(* Logix 5000 project; controller FV vendor 1 type 14 code 217 rev 31.11; software revision 31.00; part 33 of 63 *)
(* tags used below, declared in another part *)
   Alarm_Reset : BOOL;
   CheckTimeMask : INT;
   CLOCK_system_set : BOOL;
   CLOCKsetvalues : DINT[7];
   CurrentTime : DateTime;
   CWD : CHECKWORD_FLAGS;
   FR_data_file_value_to_move : DINT;
   FR_dow_addon_tag : DayOfWeek;
   FR_dow_timer : TIMER;
   FR_N120 : INT[265];   // YEAST CROP Yeast Cropping Main
   FR_N160 : INT[265];   // VESSEL Vessel Working Direc tory
   FR_N255 : INT[265];   // CHECKWORDS
   FR_N99 : INT[265];   // COMMENT Comment Lines
   FR_PANELESTOP : PlantItem;   // PANELESTOP
   FR_PILZ : PlantItem;   // PILZ
   FR_SFile : INT[255];   // SLC Equivalent System File, So Original Code Can Remain
   FR_T121 : TIMER[255];   // YEAST CROP
   FtoF_raw_input : REAL;
   FV_SFile : INT[255];   // SLC Equivalent System File, So Original Code Can Remain
   ItoF_raw_input : INT;
   One_Second_One_Scan : ALIAS FOR One_Second_1_scan;
   scale_analog_int : DINT;
   scale_analog_result : REAL;
   scale_eu_max : REAL;
   scale_eu_min : REAL;
   scale_raw_input : REAL;
   scale_raw_max : REAL;
   scale_raw_min : REAL;
   scale_routine_active : BOOL;
   scale_temp : REAL;
(* FR_Common, continued *)

ROUTINE FR_YEAST_ST_120   (* ladder *)
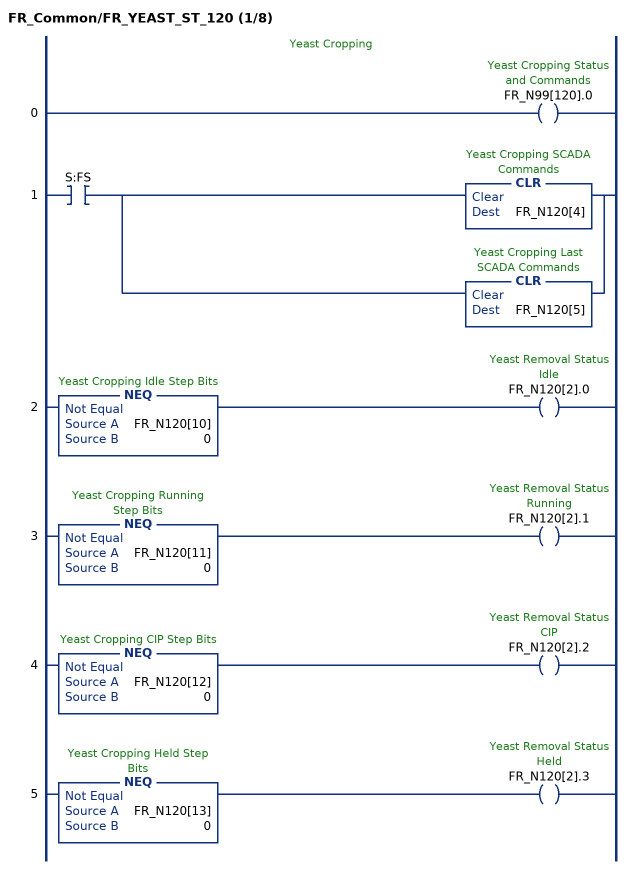
   // Yeast Cropping
   0: OTE(FR_N99[120].0);
   1: XIC(S:FS)[CLR(FR_N120[4]) ,CLR(FR_N120[5]) ];
   2: NEQ(FR_N120[10],0)OTE(FR_N120[2].0);
   3: NEQ(FR_N120[11],0)OTE(FR_N120[2].1);
   4: NEQ(FR_N120[12],0)OTE(FR_N120[2].2);
   5: NEQ(FR_N120[13],0)OTE(FR_N120[2].3);
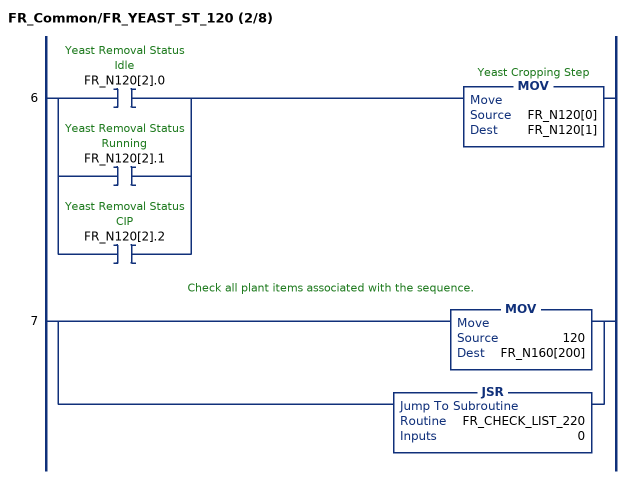
   6: [XIC(FR_N120[2].0) ,XIC(FR_N120[2].1) ,XIC(FR_N120[2].2) ]MOV(FR_N120[0],FR_N120[1]);
   // Check all plant items associated with the sequence.
   7: [MOV(120,FR_N160[200]) ,JSR(FR_CHECK_LIST_220,0) ];
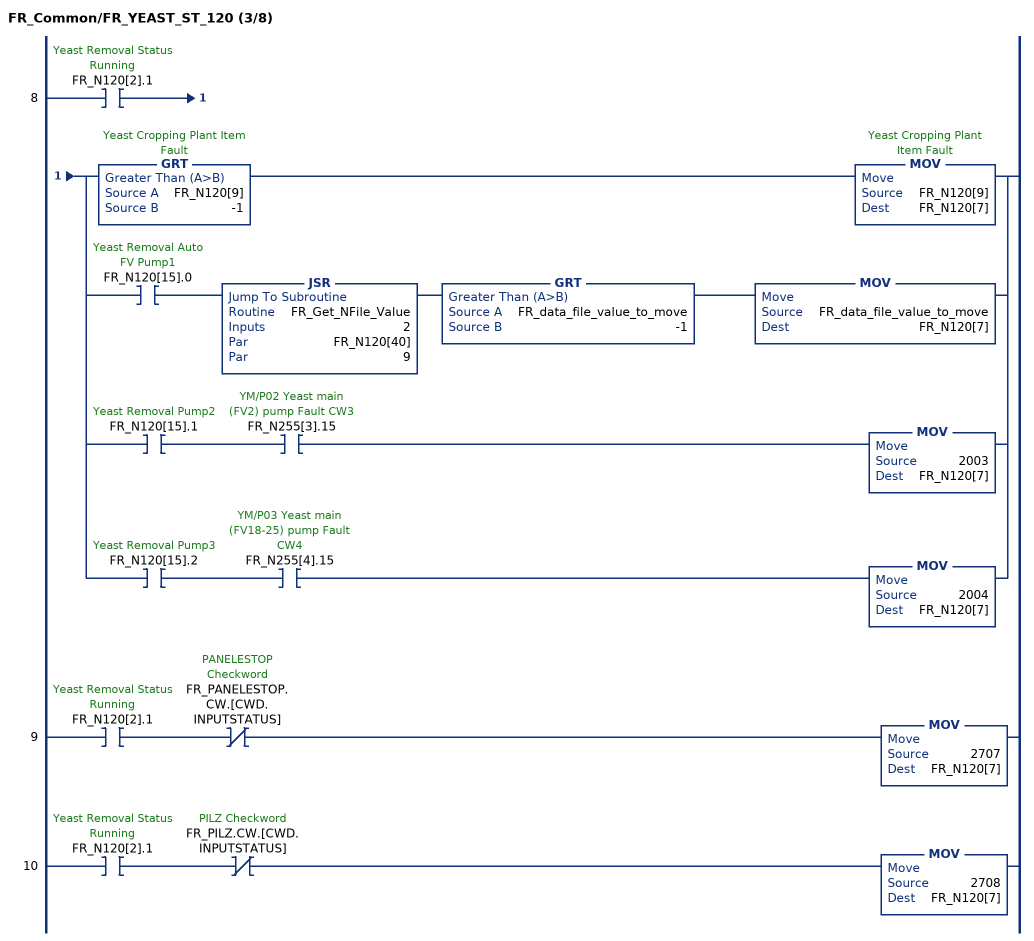
   8: XIC(FR_N120[2].1)[GRT(FR_N120[9],-1) MOV(FR_N120[9],FR_N120[7]) ,XIC(FR_N120[15].0) JSR(FR_Get_NFile_Value,2,FR_N120[40],9) GRT(FR_data_file_value_to_move,-1) MOV(FR_data_file_value_to_move,FR_N120[7]) ,XIC(FR_N120[15].1) XIC(FR_N255[3].15) MOV(2003,FR_N120[7]) ,XIC(FR_N120[15].2) XIC(FR_N255[4].15) MOV(2004,FR_N120[7]) ];
   9: XIC(FR_N120[2].1)XIO(FR_PANELESTOP.CW.[CWD.INPUTSTATUS])MOV(2707,FR_N120[7]);
   10: XIC(FR_N120[2].1)XIO(FR_PILZ.CW.[CWD.INPUTSTATUS])MOV(2708,FR_N120[7]);
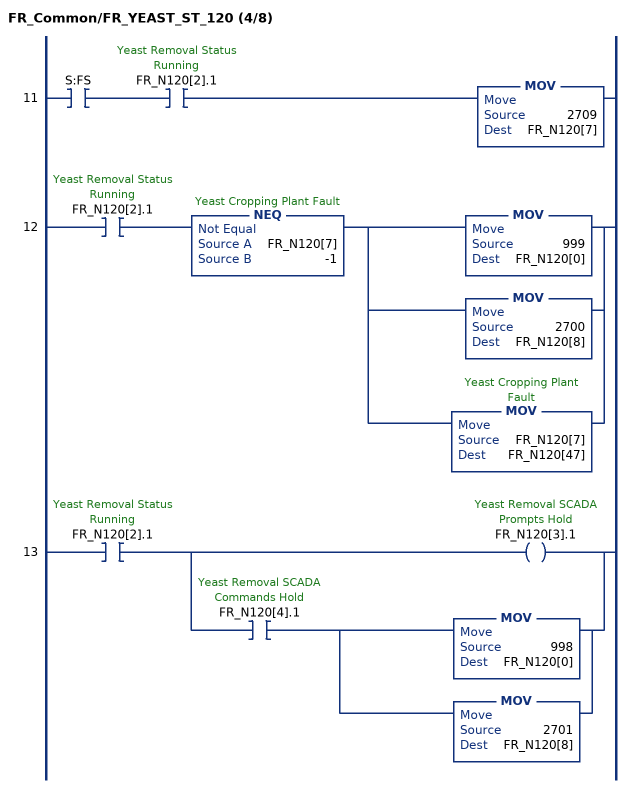
   11: XIC(S:FS)XIC(FR_N120[2].1)MOV(2709,FR_N120[7]);
   12: XIC(FR_N120[2].1)NEQ(FR_N120[7],-1)[MOV(999,FR_N120[0]) ,MOV(2700,FR_N120[8]) ,MOV(FR_N120[7],FR_N120[47]) ];
   13: XIC(FR_N120[2].1)[OTE(FR_N120[3].1) ,XIC(FR_N120[4].1) [MOV(998,FR_N120[0]) ,MOV(2701,FR_N120[8]) ] ];
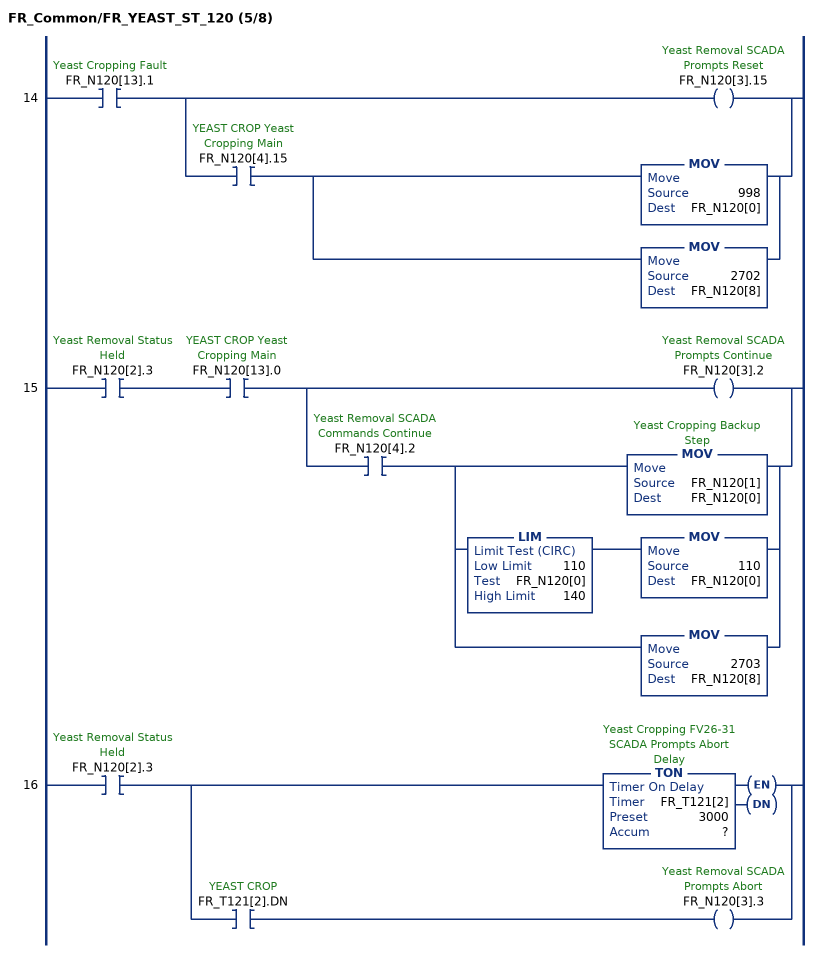
   14: XIC(FR_N120[13].1)[OTE(FR_N120[3].15) ,XIC(FR_N120[4].15) [MOV(998,FR_N120[0]) ,MOV(2702,FR_N120[8]) ] ];
   15: XIC(FR_N120[2].3)XIC(FR_N120[13].0)[OTE(FR_N120[3].2) ,XIC(FR_N120[4].2) [MOV(FR_N120[1],FR_N120[0]) ,LIM(110,FR_N120[0],140) MOV(110,FR_N120[0]) ,MOV(2703,FR_N120[8]) ] ];
   16: XIC(FR_N120[2].3)[TON(FR_T121[2],?,?) ,XIC(FR_T121[2].DN) OTE(FR_N120[3].3) ];
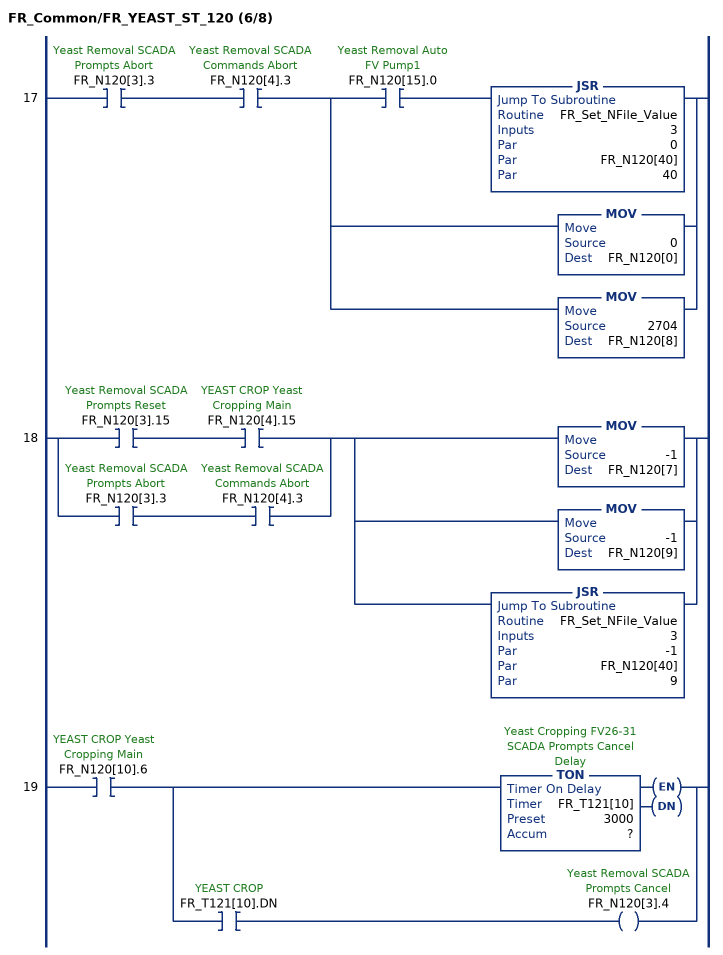
   17: XIC(FR_N120[3].3)XIC(FR_N120[4].3)[XIC(FR_N120[15].0) JSR(FR_Set_NFile_Value,3,0,FR_N120[40],40) ,MOV(0,FR_N120[0]) ,MOV(2704,FR_N120[8]) ];
   18: [XIC(FR_N120[3].15) XIC(FR_N120[4].15) ,XIC(FR_N120[3].3) XIC(FR_N120[4].3) ][MOV(-1,FR_N120[7]) ,MOV(-1,FR_N120[9]) ,JSR(FR_Set_NFile_Value,3,-1,FR_N120[40],9) ];
   19: XIC(FR_N120[10].6)[TON(FR_T121[10],?,?) ,XIC(FR_T121[10].DN) OTE(FR_N120[3].4) ];
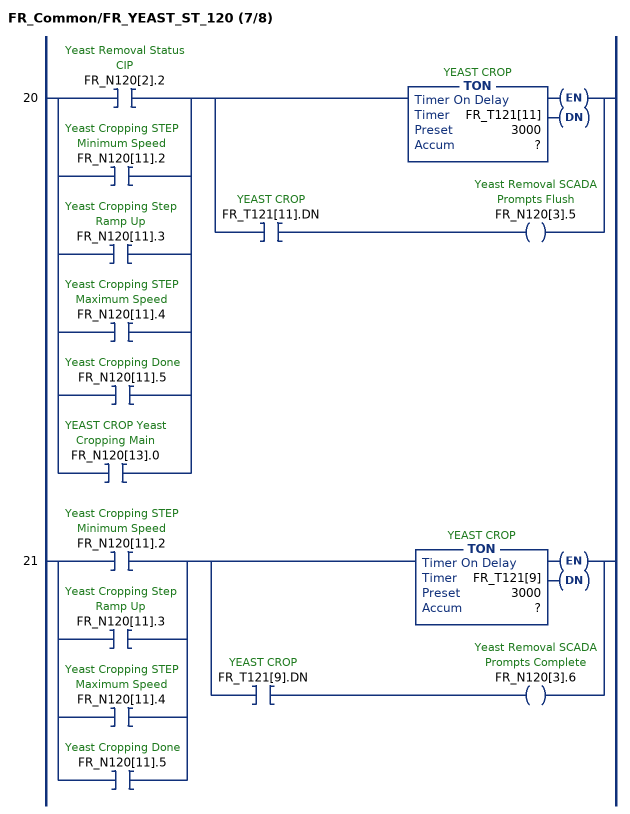
   20: [XIC(FR_N120[2].2) ,XIC(FR_N120[11].2) ,XIC(FR_N120[11].3) ,XIC(FR_N120[11].4) ,XIC(FR_N120[11].5) ,XIC(FR_N120[13].0) ][TON(FR_T121[11],?,?) ,XIC(FR_T121[11].DN) OTE(FR_N120[3].5) ];
   21: [XIC(FR_N120[11].2) ,XIC(FR_N120[11].3) ,XIC(FR_N120[11].4) ,XIC(FR_N120[11].5) ][TON(FR_T121[9],?,?) ,XIC(FR_T121[9].DN) OTE(FR_N120[3].6) ];
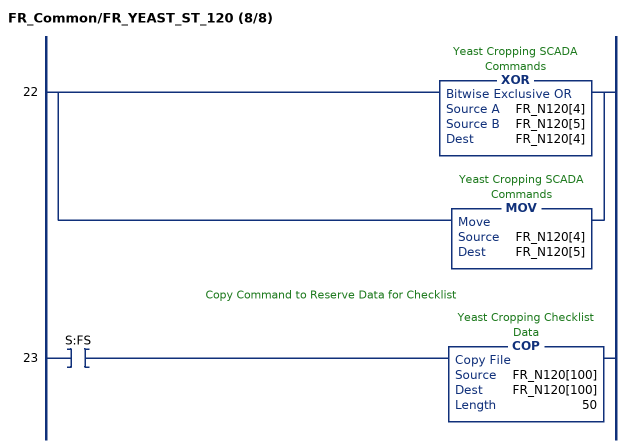
   22: [XOR(FR_N120[4],FR_N120[5],FR_N120[4]) ,MOV(FR_N120[4],FR_N120[5]) ];
   // Copy Command to Reserve Data for Checklist
   23: XIC(S:FS)COP(FR_N120[100],FR_N120[100],50);
END_ROUTINE

ROUTINE MainRoutine   (* ladder *)
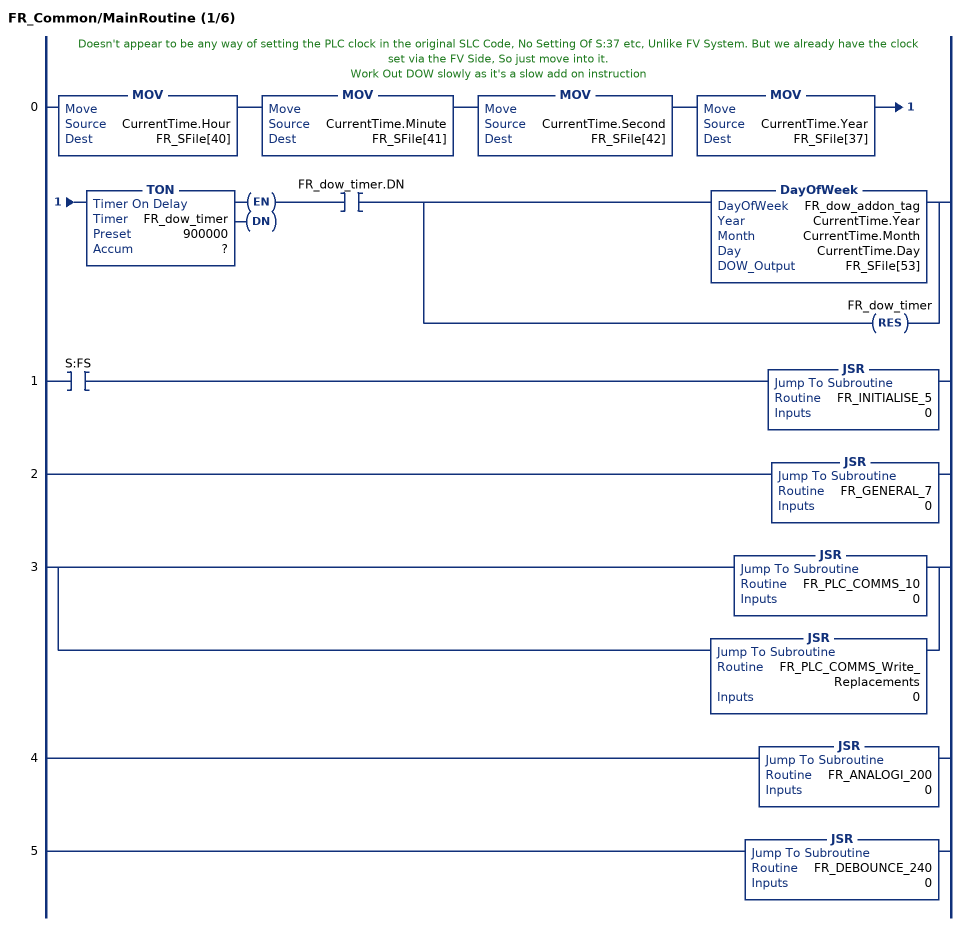
   // Doesn't appear to be any way of setting the PLC clock in the original SLC Code, No Setting Of S:37 etc, Unlike FV System. But we already have the clock set via the FV Side, So just move into it.
   // Work Out DOW slowly as it's a slow add on instruction
   0: MOV(CurrentTime.Hour,FR_SFile[40])MOV(CurrentTime.Minute,FR_SFile[41])MOV(CurrentTime.Second,FR_SFile[42])MOV(CurrentTime.Year,FR_SFile[37])TON(FR_dow_timer,?,?)XIC(FR_dow_timer.DN)[DayOfWeek(FR_dow_addon_tag,CurrentTime.Year,CurrentTime.Month,CurrentTime.Day,FR_SFile[53]) ,RES(FR_dow_timer) ];
   1: XIC(S:FS)JSR(FR_INITIALISE_5,0);
   2: JSR(FR_GENERAL_7,0);
   3: [JSR(FR_PLC_COMMS_10,0) ,JSR(FR_PLC_COMMS_Write_Replacements,0) ];
   4: JSR(FR_ANALOGI_200,0);
   5: JSR(FR_DEBOUNCE_240,0);
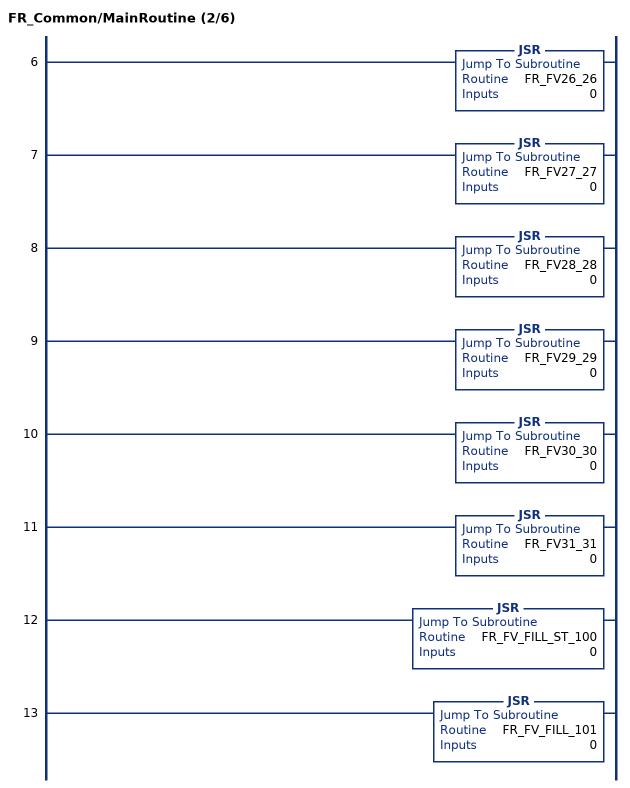
   6: JSR(FR_FV26_26,0);
   7: JSR(FR_FV27_27,0);
   8: JSR(FR_FV28_28,0);
   9: JSR(FR_FV29_29,0);
   10: JSR(FR_FV30_30,0);
   11: JSR(FR_FV31_31,0);
   12: JSR(FR_FV_FILL_ST_100,0);
   13: JSR(FR_FV_FILL_101,0);
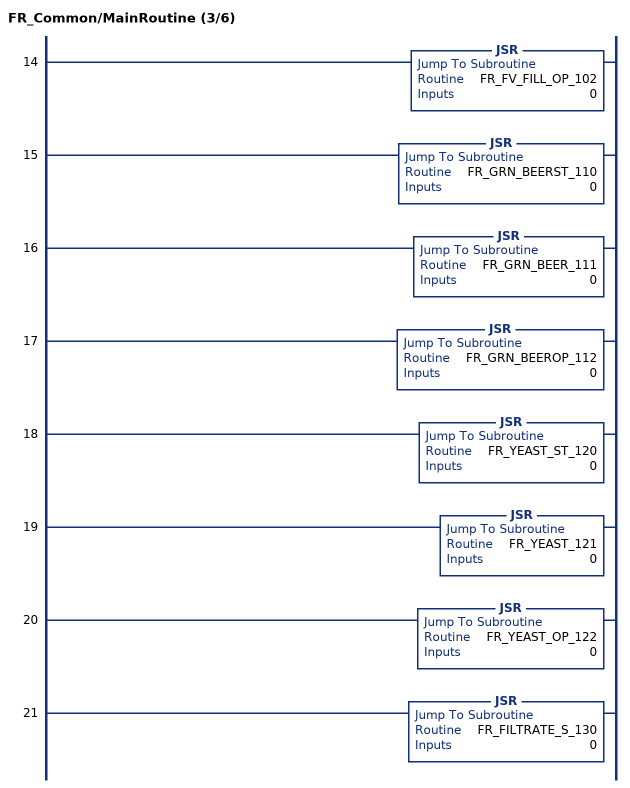
   14: JSR(FR_FV_FILL_OP_102,0);
   15: JSR(FR_GRN_BEERST_110,0);
   16: JSR(FR_GRN_BEER_111,0);
   17: JSR(FR_GRN_BEEROP_112,0);
   18: JSR(FR_YEAST_ST_120,0);
   19: JSR(FR_YEAST_121,0);
   20: JSR(FR_YEAST_OP_122,0);
   21: JSR(FR_FILTRATE_S_130,0);
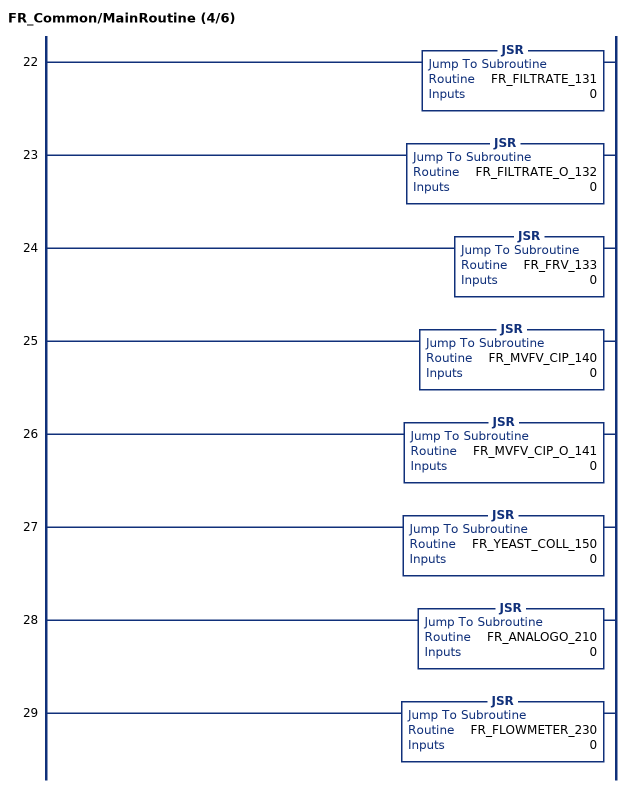
   22: JSR(FR_FILTRATE_131,0);
   23: JSR(FR_FILTRATE_O_132,0);
   24: JSR(FR_FRV_133,0);
   25: JSR(FR_MVFV_CIP_140,0);
   26: JSR(FR_MVFV_CIP_O_141,0);
   27: JSR(FR_YEAST_COLL_150,0);
   28: JSR(FR_ANALOGO_210,0);
   29: JSR(FR_FLOWMETER_230,0);
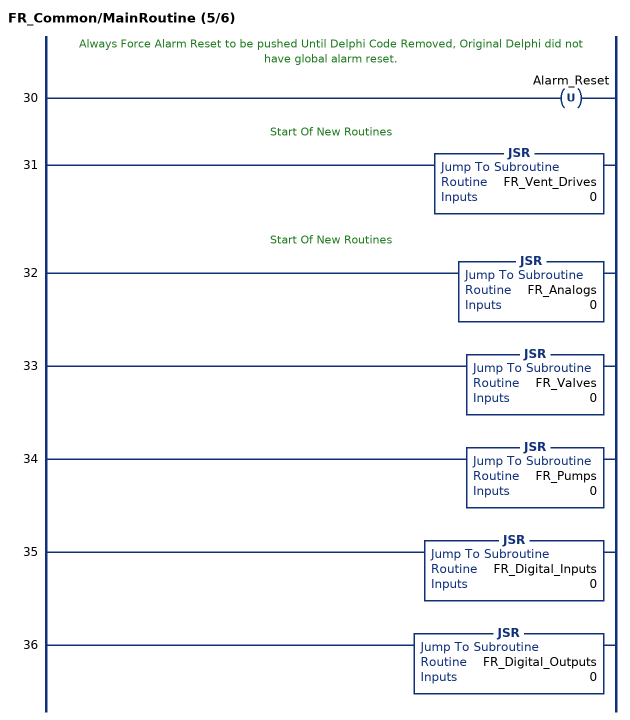
   // Always Force Alarm Reset to be pushed Until Delphi Code Removed, Original Delphi did not have global alarm reset.
   30: OTU(Alarm_Reset);
   // Start Of New Routines
   31: JSR(FR_Vent_Drives,0);
   // Start Of New Routines
   32: JSR(FR_Analogs,0);
   33: JSR(FR_Valves,0);
   34: JSR(FR_Pumps,0);
   35: JSR(FR_Digital_Inputs,0);
   36: JSR(FR_Digital_Outputs,0);
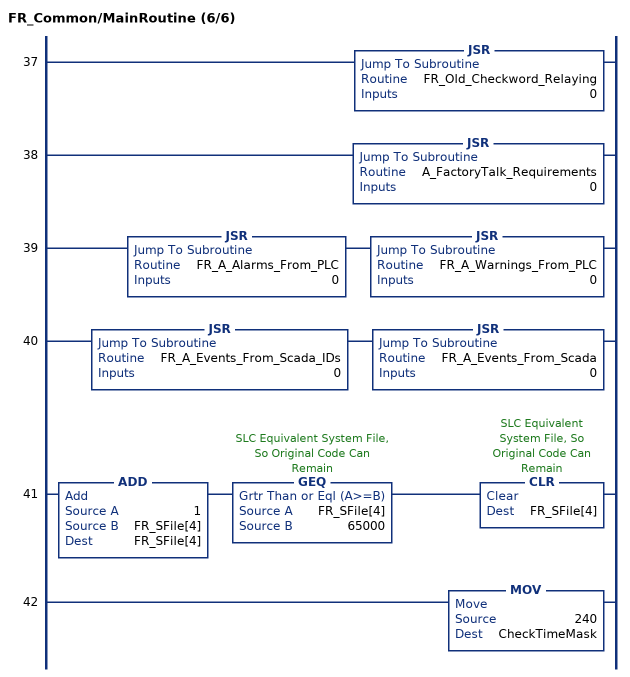
   37: JSR(FR_Old_Checkword_Relaying,0);
   38: JSR(A_FactoryTalk_Requirements,0);
   39: JSR(FR_A_Alarms_From_PLC,0)JSR(FR_A_Warnings_From_PLC,0);
   40: JSR(FR_A_Events_From_Scada_IDs,0)JSR(FR_A_Events_From_Scada,0);
   41: ADD(1,FR_SFile[4],FR_SFile[4])GEQ(FR_SFile[4],65000)CLR(FR_SFile[4]);
   42: MOV(240,CheckTimeMask);
END_ROUTINE
END_PROGRAM

PROGRAM FV_Common   (* main routine MainRoutine *)

ROUTINE A_FactoryTalk_Requirements   (* ladder *)
END_ROUTINE

ROUTINE Analog_scale_ftof   (* ladder *)
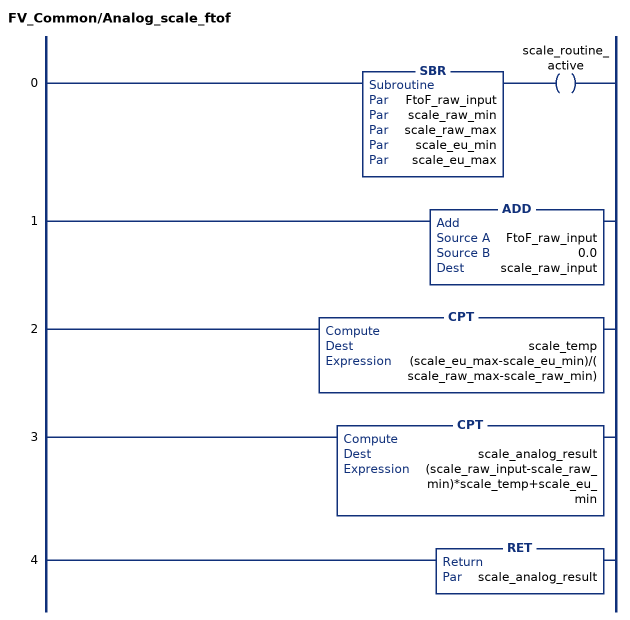
   0: SBR(FtoF_raw_input,scale_raw_min,scale_raw_max,scale_eu_min,scale_eu_max)OTE(scale_routine_active);
   1: ADD(FtoF_raw_input,0.0,scale_raw_input);
   2: CPT(scale_temp,(scale_eu_max-scale_eu_min)/(scale_raw_max-scale_raw_min));
   3: CPT(scale_analog_result,(scale_raw_input-scale_raw_min)*scale_temp+scale_eu_min);
   4: RET(scale_analog_result);
END_ROUTINE

ROUTINE Analog_Scale_FtoI   (* ladder *)
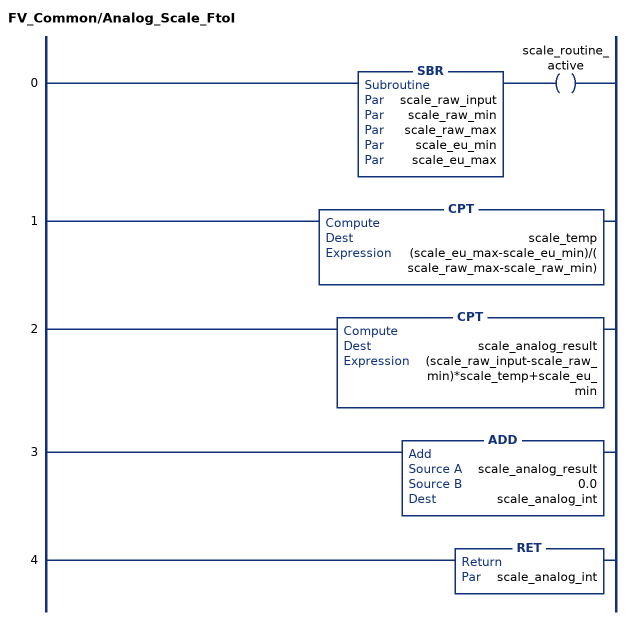
   0: SBR(scale_raw_input,scale_raw_min,scale_raw_max,scale_eu_min,scale_eu_max)OTE(scale_routine_active);
   1: CPT(scale_temp,(scale_eu_max-scale_eu_min)/(scale_raw_max-scale_raw_min));
   2: CPT(scale_analog_result,(scale_raw_input-scale_raw_min)*scale_temp+scale_eu_min);
   3: ADD(scale_analog_result,0.0,scale_analog_int);
   4: RET(scale_analog_int);
END_ROUTINE

ROUTINE Analog_Scale_ItoF   (* ladder *)
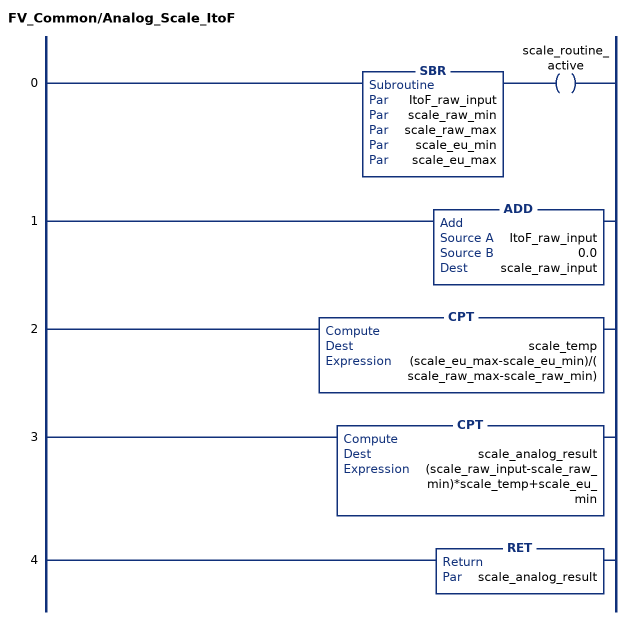
   0: SBR(ItoF_raw_input,scale_raw_min,scale_raw_max,scale_eu_min,scale_eu_max)OTE(scale_routine_active);
   1: ADD(ItoF_raw_input,0.0,scale_raw_input);
   2: CPT(scale_temp,(scale_eu_max-scale_eu_min)/(scale_raw_max-scale_raw_min));
   3: CPT(scale_analog_result,(scale_raw_input-scale_raw_min)*scale_temp+scale_eu_min);
   4: RET(scale_analog_result);
END_ROUTINE

ROUTINE ClockRoutines   (* ladder *)
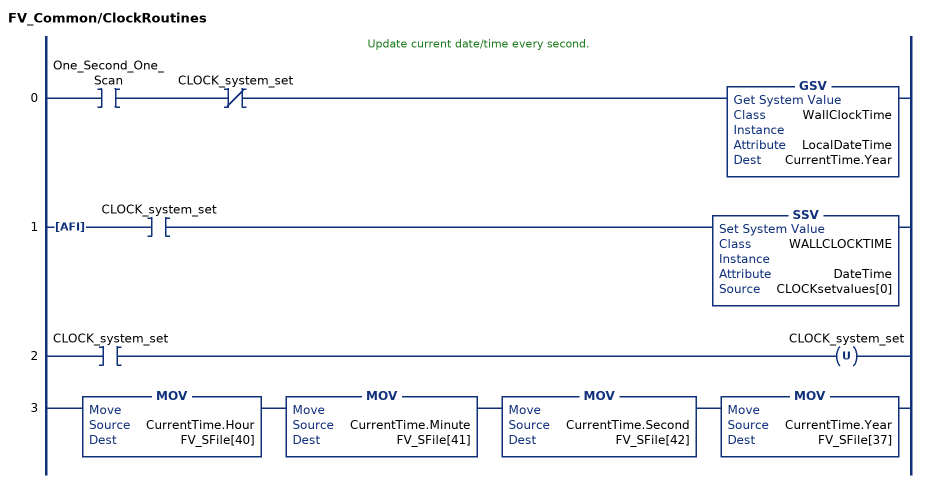
   // Update current date/time every second.
   0: XIC(One_Second_One_Scan)XIO(CLOCK_system_set)GSV(WallClockTime,,LocalDateTime,CurrentTime.Year);
   1: AFI()XIC(CLOCK_system_set)SSV(WALLCLOCKTIME,,DateTime,CLOCKsetvalues[0]);
   2: XIC(CLOCK_system_set)OTU(CLOCK_system_set);
   3: MOV(CurrentTime.Hour,FV_SFile[40])MOV(CurrentTime.Minute,FV_SFile[41])MOV(CurrentTime.Second,FV_SFile[42])MOV(CurrentTime.Year,FV_SFile[37]);
END_ROUTINE
